Fault WB1[30].25'; 986 '~S001R03 Sealer Ctrlr 2 Required Rezeroing WB1[30].26'; 987 '~S001R03 Mig Barrel Replacement Warning WB1[30].27'; 988 '~S001R03 Mig Barrel Replacement Required WB1[30].28'; 989 '~S001R03 In Touch Up Mode WB1[30].29'; 990 '~S001R03 Touch Up Mode Not Enabled WB1[30].30'; 991 '~Spare WB1[30].31'; 992 '~S001R03 Laser Controller Fault WB1[31].0'; 993 '~S001R03 Laser Dirty Glass Warning WB1[31].1'; 994 '~S001R03 Laser Warning WB1[31].2'; 995 '~Spare WB1[31].3'; 996 '~Spare WB1[31].4'; 997 '~Spare WB1[31].5'; 998 '~Spare WB1[31].6'; 999 '~Spare WB1[31].7'; 1000 '~Spare WB1[31].8'; 1001 '~Spare WB1[31].9'; 1002 '~Spare WB1[31].10'; 1003 '~Spare WB1[31].11'; 1004 '~Spare WB1[31].12'; 1005 '~Spare WB1[31].13'; 1006 '~Spare WB1[31].14'; 1007 '~Spare WB1[31].15'; 1008 '~Spare WB1[31].16'; 1009 '~Spare WB1[31].17'; 1010 '~Spare WB1[31].18'; 1011 '~Spare WB1[31].19'; 1012 '~Spare WB1[31].20'; 1013 '~Spare WB1[31].21'; 1014 '~Spare WB1[31].22'; 1015 '~Spare WB1[31].23'; 1016 '~Spare WB1[31].24'; 1017 '~Spare WB1[31].25'; 1018 '~Spare WB1[31].26'; 1019 '~Spare WB1[31].27'; 1020 '~Spare WB1[31].28'; 1021 '~Spare WB1[31].29'; 1022 '~Spare WB1[31].30'; 1023 '~Spare WB1[31].31'; 1024 '~Spare WB1[32].0'; 1025 '~Spare WB1[32].1'; 1026 '~Spare WB1[32].2'; 1027 '~Spare WB1[32].3'; 1028 '~Spare WB1[32].4'; 1029 '~Spare WB1[32].5'; 1030 '~Spare WB1[32].6'; 1031 '~Spare WB1[32].7'; 1032 '~Spare WB1[32].8'; 1033 '~Spare WB1[32].9'; 1034 '~Spare WB1[32].10'; 1035 '~Spare WB1[32].11'; 1036 '~Spare WB1[32].12'; 1037 '~Spare WB1[32].13'; 1038 '~Spare WB1[32].14'; 1039 '~Spare WB1[32].15'; 1040 '~Spare WB1[32].16'; 1041 '~Spare WB1[32].17'; 1042 '~Spare WB1[32].18'; 1043 '~Spare WB1[32].19'; 1044 '~Spare WB1[32].20'; 1045 '~Spare WB1[32].21'; 1046 '~Spare WB1[32].22'; 1047 '~Spare WB1[32].23'; 1048 '~Spare WB1[32].24'; 1049 '~Spare WB1[32].25'; 1050 '~Spare WB1[32].26'; 1051 '~Spare WB1[32].27'; 1052 '~Spare WB1[32].28'; 1053 '~Spare WB1[32].29'; 1054 '~Spare WB1[32].30'; 1055 '~Spare WB1[32].31'; 1056 '~Spare WB1[33].0'; 1057 '~Spare WB1[33].1'; 1058 '~Spare WB1[33].2'; 1059 '~Spare WB1[33].3'; 1060 '~Spare WB1[33].4'; 1061 '~Spare WB1[33].5'; 1062 '~Spare WB1[33].6'; 1063 '~Spare WB1[33].7'; 1064 '~Spare WB1[33].8'; 1065 '~Spare WB1[33].9'; 1066 '~Spare WB1[33].10'; 1067 '~Spare WB1[33].11'; 1068 '~Spare WB1[33].12'; 1069 '~Spare WB1[33].13'; 1070 '~Spare WB1[33].14'; 1071 '~Spare WB1[33].15'; 1072 '~Spare WB1[33].16'; 1073 '~Spare WB1[33].17'; 1074 '~Spare WB1[33].18'; 1075 '~Spare WB1[33].19'; 1076 '~Spare WB1[33].20'; 1077 '~Spare WB1[33].21'; 1078 '~Spare WB1[33].22'; 1079 '~Spare WB1[33].23'; 1080 '~Spare WB1[33].24'; 1081 '~Spare WB1[33].25'; 1082 '~Spare WB1[33].26'; 1083 '~Spare WB1[33].27'; 1084 '~Spare WB1[33].28'; 1085 '~Spare WB1[33].29'; 1086 '~Spare WB1[33].30'; 1087 '~Spare WB1[33].31'; 1088 '~S001R04 Waiting Zone #1 Not Clear WB1[34].0'; 1089 '~S001R04 Waiting Zone #2 Not Clear WB1[34].1'; 1090 '~S001R04 Waiting Zone #3 Not Clear WB1[34].2'; 1091 '~S001R04 Waiting Zone #4 Not Clear WB1[34].3'; 1092 '~S001R04 Waiting Zone #5 Not Clear WB1[34].4'; 1093 '~S001R04 Waiting Zone #6 Not Clear WB1[34].5'; 1094 '~S001R04 Waiting Zone #7 Not Clear WB1[34].6'; 1095 '~S001R04 Waiting Zone #8 Not Clear WB1[34].7'; 1096 '~S001R04 Waiting Zone #9 Not Clear WB1[34].8'; 1097 '~S001R04 Waiting Zone #10 Not Clear WB1[34].9'; 1098 '~S001R04 Waiting Zone #11 Not Clear WB1[34].10'; 1099 '~S001R04 Waiting Zone #12 Not Clear WB1[34].11'; 1100 '~S001R04 Waiting Zone #13 Not Clear WB1[34].12'; 1101 '~S001R04 Waiting Zone #14 Not Clear WB1[34].13'; 1102 '~S001R04 Waiting Tip Dress Zone #1 Not Clear WB1[34].14'; 1103 '~S001R04 Waiting Tip Dress Zone #2 Not Clear WB1[34].15'; 1104 '~S001R04 Adjacent Robot xx-xx In Teach WB1[34].16'; 1105 '~S001R04 Adjacent Robot xx-xx In Teach WB1[34].17'; 1106 '~S001R04 Adjacent Robot xx-xx In Teach WB1[34].18'; 1107 '~S001R04 Adjacent Robot xx-xx In Teach WB1[34].19'; 1108 '~S001R04 Adjacent Robot xx-xx In Teach WB1[34].20'; 1109 '~S001R04 Adjacent Robot xx-xx In Teach WB1[34].21'; 1110 '~S001R04 Adjacent Robot xx-xx In Teach WB1[34].22'; 1111 '~S001R04 Adjacent Robot xx-xx In Teach WB1[34].23'; 1112 '~S001R04 Adjacent Robot xx-xx In Teach WB1[34].24'; 1113 '~S001R04 Adjacent Robot xx-xx In Teach WB1[34].25'; 1114 '~Spare WB1[34].26'; 1115 '~Spare WB1[34].27'; 1116 '~Spare WB1[34].28'; 1117 '~S001R04 Robot Not Clear Of Fixture WB1[34].29'; 1118 '~Spare WB1[34].30'; 1119 '~Spare WB1[34].31'; 1120 '~Spare WB1[35].0'; 1121 '~Spare WB1[35].1'; 1122 '~Spare WB1[35].2'; 1123 '~Spare WB1[35].3'; 1124 '~Spare WB1[35].4'; 1125 '~Spare WB1[35].5'; 1126 '~Spare WB1[35].6'; 1127 '~Spare WB1[35].7'; 1128 '~Spare WB1[35].8'; 1129 '~Spare WB1[35].9'; 1130 '~Spare WB1[35].10'; 1131 '~Spare WB1[35].11'; 1132 '~Spare WB1[35].12'; 1133 '~Spare WB1[35].13'; 1134 '~Spare WB1[35].14'; 1135 '~Spare WB1[35].15'; 1136 '~Spare WB1[35].16'; 1137 '~Spare WB1[35].17'; 1138 '~Spare WB1[35].18'; 1139 '~Spare WB1[35].19'; 1140 '~Spare WB1[35].20'; 1141 '~Spare WB1[35].21'; 1142 '~Spare WB1[35].22'; 1143 '~Spare WB1[35].23'; 1144 '~Spare WB1[35].24'; 1145 '~Spare WB1[35].25'; 1146 '~Spare WB1[35].26'; 1147 '~Spare WB1[35].27'; 1148 '~Spare WB1[35].28'; 1149 '~Spare WB1[35].29'; 1150 '~Spare WB1[35].30'; 1151 '~Spare WB1[35].31'; 1152 '~S001R04 Cycle Overtime WB1[36].0'; 1153 '~S001R04 In Bypass WB1[36].1'; 1154 '~S001R04 Battery Low WB1[36].2'; 1155 '~S001R04 Servo Over Torque WB1[36].3'; 1156 '~S001R04 Process Retry In Progress WB1[36].4'; 1157 '~Spare WB1[36].5'; 1158 '~S001R04 Robot Edit Occurred Ext App WB1[36].6'; 1159 '~S001R04 Robot Input Simmed WB1[36].7'; 1160 '~S001R04 Robot Output Simmed WB1[36].8'; 1161 '~Spare WB1[36].9'; 1162 '~Spare WB1[36].10'; 1163 '~Spare WB1[36].11'; 1164 '~Spare WB1[36].12'; 1165 '~Spare WB1[36].13'; 1166 '~Spare WB1[36].14'; 1167 '~Spare WB1[36].15'; 1168 '~S001R04F1B1.M.ModuleFlt - Externa App 1 I/O Module Warning WB1[36].16'; 1169 '~S001R04F2B1.M.ModuleFlt - Externa App 2 I/O Module Warning WB1[36].17'; 1170 '~S001R04F3B1.M.ModuleFlt - Externa App 3 I/O Module Warning WB1[36].18'; 1171 '~Spare WB1[36].19'; 1172 '~Spare WB1[36].20'; 1173 '~Spare WB1[36].21'; 1174 '~Spare WB1[36].22'; 1175 '~Spare WB1[36].23'; 1176 '~S001R04ES1 - S001R04 EtherNet Switch Port At Half Duplex WB1[36].24'; 1177 '~S001R04ES1 - S001R04 EtherNet Switch Config Changes Not Saved WB1[36].25'; 1178 '~S001R04ES1 - S001R04 EtherNet Switch Configuration Changed WB1[36].26'; 1179 '~S001R04ES1 - S001R04 EtherNet Switch Port With Excessive Errors WB1[36].27'; 1180 '~S001R04ES1 - S001R04 EtherNet Switch Port With Utilization Warning WB1[36].28'; 1181 '~S001R04ES1 - S001R04 EtherNet Switch Changes Require Reboot WB1[36].29'; 1182 '~Spare WB1[36].30'; 1183 '~Spare WB1[36].31'; 1184 '~Spare WB1[37].0'; 1185 '~Spare WB1[37].1'; 1186 '~S001R04 Servo Gun Tip Calib Request 1 WB1[37].2'; 1187 '~S001R04 I-Available Warning 1 WB1[37].3'; 1188 '~S001R04 Tip Dress Motor 1 Fault Bypassed WB1[37].4'; 1189 '~S001R04 Tip Change Notice 1 WB1[37].5'; 1190 '~S001R04 Bypass Tip Dresser 1 Selected WB1[37].6'; 1191 '~S001R04 Auto Tip Changer Low 1 WB1[37].7'; 1192 '~S001R04 Auto Tip Changer Empty 1 WB1[37].8'; 1193 '~S001R04 Tip Wear Ratio Warning 1 - Touch Up Tip Dress Program WB1[37].9'; 1194 '~S001R04 Stud Weld 1 Maintenance Reqd WB1[37].10'; 1195 '~S001R04 Stud Weld 1 Low Stud Warning WB1[37].11'; 1196 '~Spare WB1[37].12'; 1197 '~S001R04 Rivet 1 Low Rivet Warning WB1[37].13'; 1198 '~S001R04 Rivet 1 - Skip Once Initiated from Robot TP WB1[37].14'; 1199 '~S001R04 Rivet 1 - Skip Remaining Initiated from Robot TP WB1[37].15'; 1200 '~S001R04 Rivet 1 Preventive Maintenace Required WB1[37].16'; 1201 '~S001R04 Rivet 1 Magazine Low WB1[37].17'; 1202 '~S001R04 Tip Change 1 Bypassed WB1[37].18'; 1203 '~S001R04 Mig Weld Fluid Level Low WB1[37].19'; 1204 '~S001R04 Weld Ctrlr 1 Adaptive Mode Is Disabled WB1[37].20'; 1205 '~S001R04 Tip Cutter 1 Warning WB1[37].21'; 1206 '~S001R04 Rivet 1 Tape-Cut Required WB1[37].22'; 1207 '~S001R04 Wire Feeder Motor Over Current WB1[37].23'; 1208 '~Spare WB1[37].24'; 1209 '~S001R04 Sealer Ctrlr 1 Minor Fault WB1[37].25'; 1210 '~S001R04 Sealer Ctrlr 1 Required Rezeroing WB1[37].26'; 1211 '~S001R04 Loaded To Average WB1[37].27'; 1212 '~S001R04 Vision Process Aborted WB1[37].28'; 1213 '~S001R04 Vision System Trending WB1[37].29'; 1214 '~S001R04 Vision Out Of Tolerance WB1[37].30'; 1215 '~Spare WB1[37].31'; 1216 '~Spare WB1[38].0'; 1217 '~Spare WB1[38].1'; 1218 '~S001R04 Servo Gun Tip Calib Request 2 WB1[38].2'; 1219 '~S001R04 I-Available Warning 2 WB1[38].3'; 1220 '~S001R04 Tip Dress Motor 2 Fault Bypassed WB1[38].4'; 1221 '~S001R04 Tip Change Notice 2 WB1[38].5'; 1222 '~S001R04 Bypass Tip Dresser 2 Selected WB1[38].6'; 1223 '~S001R04 Auto Tip Changer Low 2 WB1[38].7'; 1224 '~S001R04 Auto Tip Changer Empty 2 WB1[38].8'; 1225 '~S001R04 Tip Wear Ratio Warning 2 - Touch Up Tip Dress Program WB1[38].9'; 1226 '~S001R04 Stud Weld 2 Maintenance Reqd WB1[38].10'; 1227 '~S001R04 Stud Weld 2 Low Stud Warning WB1[38].11'; 1228 '~Spare WB1[38].12'; 1229 '~S001R04 Rivet 2 Low Rivet Warning WB1[38].13'; 1230 '~S001R04 Rivet 2 - Skip Once Initiated from Robot TP WB1[38].14'; 1231 '~S001R04 Rivet 2 - Skip Remaining Initiated from Robot TP WB1[38].15'; 1232 '~S001R04 Rivet 2 Preventive Maintenace Required WB1[38].16'; 1233 '~S001R04 Rivet 2 Magazine Low WB1[38].17'; 1234 '~S001R04 Tip Change 2 Bypassed WB1[38].18'; 1235 '~S001R04 Laser Dirty Glass Warning WB1[38].19'; 1236 '~S001R04 Weld Ctrlr 2 Adaptive Mode Is Disabled WB1[38].20'; 1237 '~S001R04 Tip Cutter 2 Warning WB1[38].21'; 1238 '~S001R04 Rivet 2 Tape-Cut Required WB1[38].22'; 1239 '~S001R04 Mig Tip Nozzel Replacement Warning WB1[38].23'; 1240 '~S001R04 Mig Tip Nozzel Replacement Required WB1[38].24'; 1241 '~S001R04 Sealer Ctrlr 2 Minor Fault WB1[38].25'; 1242 '~S001R04 Sealer Ctrlr 2 Required Rezeroing WB1[38].26'; 1243 '~S001R04 Mig Barrel Replacement Warning WB1[38].27'; 1244 '~S001R04 Mig Barrel Replacement Required WB1[38].28'; 1245 '~S001R04 In Touch Up Mode WB1[38].29'; 1246 '~S001R04 Touch Up Mode Not Enabled WB1[38].30'; 1247 '~Spare WB1[38].31'; 1248 '~S001R04 Laser Controller Fault WB1[39].0'; 1249 '~S001R04 Laser Dirty Glass Warning WB1[39].1'; 1250 '~S001R04 Laser Warning WB1[39].2'; 1251 '~Spare WB1[39].3'; 1252 '~Spare WB1[39].4'; 1253 '~Spare WB1[39].5'; 1254 '~Spare WB1[39].6'; 1255 '~Spare WB1[39].7'; 1256 '~Spare WB1[39].8'; 1257 '~Spare WB1[39].9'; 1258 '~Spare WB1[39].10'; 1259 '~Spare WB1[39].11'; 1260 '~Spare WB1[39].12'; 1261 '~Spare WB1[39].13'; 1262 '~Spare WB1[39].14'; 1263 '~Spare WB1[39].15'; 1264 '~Spare WB1[39].16'; 1265 '~Spare WB1[39].17'; 1266 '~Spare WB1[39].18'; 1267 '~Spare WB1[39].19'; 1268 '~Spare WB1[39].20'; 1269 '~Spare WB1[39].21'; 1270 '~Spare WB1[39].22'; 1271 '~Spare WB1[39].23'; 1272 '~Spare WB1[39].24'; 1273 '~Spare WB1[39].25'; 1274 '~Spare WB1[39].26'; 1275 '~Spare WB1[39].27'; 1276 '~Spare WB1[39].28'; 1277 '~Spare WB1[39].29'; 1278 '~Spare WB1[39].30'; 1279 '~Spare WB1[39].31'; 1280 '~Spare WB1[40].0'; 1281 '~Spare WB1[40].1'; 1282 '~Spare WB1[40].2'; 1283 '~Spare WB1[40].3'; 1284 '~Spare WB1[40].4'; 1285 '~Spare WB1[40].5'; 1286 '~Spare WB1[40].6'; 1287 '~Spare WB1[40].7'; 1288 '~Spare WB1[40].8'; 1289 '~Spare WB1[40].9'; 1290 '~Spare WB1[40].10'; 1291 '~Spare WB1[40].11'; 1292 '~Spare WB1[40].12'; 1293 '~Spare WB1[40].13'; 1294 '~Spare WB1[40].14'; 1295 '~Spare WB1[40].15'; 1296 '~Spare WB1[40].16'; 1297 '~Spare WB1[40].17'; 1298 '~Spare WB1[40].18'; 1299 '~Spare WB1[40].19'; 1300 '~Spare WB1[40].20'; 1301 '~Spare WB1[40].21'; 1302 '~Spare WB1[40].22'; 1303 '~Spare WB1[40].23'; 1304 '~Spare WB1[40].24'; 1305 '~Spare WB1[40].25'; 1306 '~Spare WB1[40].26'; 1307 '~Spare WB1[40].27'; 1308 '~Spare WB1[40].28'; 1309 '~Spare WB1[40].29'; 1310 '~Spare WB1[40].30'; 1311 '~Spare WB1[40].31'; 1312 '~Spare WB1[41].0'; 1313 '~Spare WB1[41].1'; 1314 '~Spare WB1[41].2'; 1315 '~Spare WB1[41].3'; 1316 '~Spare WB1[41].4'; 1317 '~Spare WB1[41].5'; 1318 '~Spare WB1[41].6'; 1319 '~Spare WB1[41].7'; 1320 '~Spare WB1[41].8'; 1321 '~Spare WB1[41].9'; 1322 '~Spare WB1[41].10'; 1323 '~Spare WB1[41].11'; 1324 '~Spare WB1[41].12'; 1325 '~Spare WB1[41].13'; 1326 '~Spare WB1[41].14'; 1327 '~Spare WB1[41].15'; 1328 '~Spare WB1[41].16'; 1329 '~Spare WB1[41].17'; 1330 '~Spare WB1[41].18'; 1331 '~Spare WB1[41].19'; 1332 '~Spare WB1[41].20'; 1333 '~Spare WB1[41].21'; 1334 '~Spare WB1[41].22'; 1335 '~Spare WB1[41].23'; 1336 '~Spare WB1[41].24'; 1337 '~Spare WB1[41].25'; 1338 '~Spare WB1[41].26'; 1339 '~Spare WB1[41].27'; 1340 '~Spare WB1[41].28'; 1341 '~Spare WB1[41].29'; 1342 '~Spare WB1[41].30'; 1343 '~Spare WB1[41].31'; 1344 '~S001R05 Waiting Zone #1 Not Clear WB1[42].0'; 1345 '~S001R05 Waiting Zone #2 Not Clear WB1[42].1'; 1346 '~S001R05 Waiting Zone #3 Not Clear WB1[42].2'; 1347 '~S001R05 Waiting Zone #4 Not Clear WB1[42].3'; 1348 '~S001R05 Waiting Zone #5 Not Clear WB1[42].4'; 1349 '~S001R05 Waiting Zone #6 Not Clear WB1[42].5'; 1350 '~S001R05 Waiting Zone #7 Not Clear WB1[42].6'; 1351 '~S001R05 Waiting Zone #8 Not Clear WB1[42].7'; 1352 '~S001R05 Waiting Zone #9 Not Clear WB1[42].8'; 1353 '~S001R05 Waiting Zone #10 Not Clear WB1[42].9'; 1354 '~S001R05 Waiting Zone #11 Not Clear WB1[42].10'; 1355 '~S001R05 Waiting Zone #12 Not Clear WB1[42].11'; 1356 '~S001R05 Waiting Zone #13 Not Clear WB1[42].12'; 1357 '~S001R05 Waiting Zone #14 Not Clear WB1[42].13'; 1358 '~S001R05 Waiting Tip Dress Zone #1 Not Clear WB1[42].14'; 1359 '~S001R05 Waiting Tip Dress Zone #2 Not Clear WB1[42].15'; 1360 '~S001R05 Adjacent Robot xx-xx In Teach WB1[42].16'; 1361 '~S001R05 Adjacent Robot xx-xx In Teach WB1[42].17'; 1362 '~S001R05 Adjacent Robot xx-xx In Teach WB1[42].18'; 1363 '~S001R05 Adjacent Robot xx-xx In Teach WB1[42].19'; 1364 '~S001R05 Adjacent Robot xx-xx In Teach WB1[42].20'; 1365 '~S001R05 Adjacent Robot xx-xx In Teach WB1[42].21'; 1366 '~S001R05 Adjacent Robot xx-xx In Teach WB1[42].22'; 1367 '~S001R05 Adjacent Robot xx-xx In Teach WB1[42].23'; 1368 '~S001R05 Adjacent Robot xx-xx In Teach WB1[42].24'; 1369 '~S001R05 Adjacent Robot xx-xx In Teach WB1[42].25'; 1370 '~Spare WB1[42].26'; 1371 '~Spare WB1[42].27'; 1372 '~Spare WB1[42].28'; 1373 '~S001R05 Robot Not Clear Of Fixture WB1[42].29'; 1374 '~Spare WB1[42].30'; 1375 '~Spare WB1[42].31'; 1376 '~Spare WB1[43].0'; 1377 '~Spare WB1[43].1'; 1378 '~Spare WB1[43].2'; 1379 '~Spare WB1[43].3'; 1380 '~Spare WB1[43].4'; 1381 '~Spare WB1[43].5'; 1382 '~Spare WB1[43].6'; 1383 '~Spare WB1[43].7'; 1384 '~Spare WB1[43].8'; 1385 '~Spare WB1[43].9'; 1386 '~Spare WB1[43].10'; 1387 '~Spare WB1[43].11'; 1388 '~Spare WB1[43].12'; 1389 '~Spare WB1[43].13'; 1390 '~Spare WB1[43].14'; 1391 '~Spare WB1[43].15'; 1392 '~Spare WB1[43].16'; 1393 '~Spare WB1[43].17'; 1394 '~Spare WB1[43].18'; 1395 '~Spare WB1[43].19'; 1396 '~Spare WB1[43].20'; 1397 '~Spare WB1[43].21'; 1398 '~Spare WB1[43].22'; 1399 '~Spare WB1[43].23'; 1400 '~Spare WB1[43].24'; 1401 '~Spare WB1[43].25'; 1402 '~Spare WB1[43].26'; 1403 '~Spare WB1[43].27'; 1404 '~Spare WB1[43].28'; 1405 '~Spare WB1[43].29'; 1406 '~Spare WB1[43].30'; 1407 '~Spare WB1[43].31'; 1408 '~S001R05 Cycle Overtime WB1[44].0'; 1409 '~S001R05 In Bypass WB1[44].1'; 1410 '~S001R05 Battery Low WB1[44].2'; 1411 '~S001R05 Servo Over Torque WB1[44].3'; 1412 '~S001R05 Process Retry In Progress WB1[44].4'; 1413 '~Spare WB1[44].5'; 1414 '~S001R05 Robot Edit Occurred Ext App WB1[44].6'; 1415 '~S001R05 Robot Input Simmed WB1[44].7'; 1416 '~S001R05 Robot Output Simmed WB1[44].8'; 1417 '~Spare WB1[44].9'; 1418 '~Spare WB1[44].10'; 1419 '~Spare WB1[44].11'; 1420 '~Spare WB1[44].12'; 1421 '~Spare WB1[44].13'; 1422 '~Spare WB1[44].14'; 1423 '~Spare WB1[44].15'; 1424 '~S001R05F1B1.M.ModuleFlt - Externa App 1 I/O Module Warning WB1[44].16'; 1425 '~S001R05F2B1.M.ModuleFlt - Externa App 2 I/O Module Warning WB1[44].17'; 1426 '~S001R05F3B1.M.ModuleFlt - Externa App 3 I/O Module Warning WB1[44].18'; 1427 '~Spare WB1[44].19'; 1428 '~Spare WB1[44].20'; 1429 '~Spare WB1[44].21'; 1430 '~Spare WB1[44].22'; 1431 '~Spare WB1[44].23'; 1432 '~S001R05ES1 - S001R05 EtherNet Switch Port At Half Duplex WB1[44].24'; 1433 '~S001R05ES1 - S001R05 EtherNet Switch Config Changes Not Saved WB1[44].25'; 1434 '~S001R05ES1 - S001R05 EtherNet Switch Configuration Changed WB1[44].26'; 1435 '~S001R05ES1 - S001R05 EtherNet Switch Port With Excessive Errors WB1[44].27'; 1436 '~S001R05ES1 - S001R05 EtherNet Switch Port With Utilization Warning WB1[44].28'; 1437 '~S001R05ES1 - S001R05 EtherNet Switch Changes Require Reboot WB1[44].29'; 1438 '~Spare WB1[44].30'; 1439 '~Spare WB1[44].31'; 1440 '~Spare WB1[45].0'; 1441 '~Spare WB1[45].1'; 1442 '~S001R05 Servo Gun Tip Calib Request 1 WB1[45].2'; 1443 '~S001R05 I-Available Warning 1 WB1[45].3'; 1444 '~S001R05 Tip Dress Motor 1 Fault Bypassed WB1[45].4'; 1445 '~S001R05 Tip Change Notice 1 WB1[45].5'; 1446 '~S001R05 Bypass Tip Dresser 1 Selected WB1[45].6'; 1447 '~S001R05 Auto Tip Changer Low 1 WB1[45].7'; 1448 '~S001R05 Auto Tip Changer Empty 1 WB1[45].8'; 1449 '~S001R05 Tip Wear Ratio Warning 1 - Touch Up Tip Dress Program WB1[45].9'; 1450 '~S001R05 Stud Weld 1 Maintenance Reqd WB1[45].10'; 1451 '~S001R05 Stud Weld 1 Low Stud Warning WB1[45].11'; 1452 '~Spare WB1[45].12'; 1453 '~S001R05 Rivet 1 Low Rivet Warning WB1[45].13'; 1454 '~S001R05 Rivet 1 - Skip Once Initiated from Robot TP WB1[45].14'; 1455 '~S001R05 Rivet 1 - Skip Remaining Initiated from Robot TP WB1[45].15'; 1456 '~S001R05 Rivet 1 Preventive Maintenace Required WB1[45].16'; 1457 '~S001R05 Rivet 1 Magazine Low WB1[45].17'; 1458 '~S001R05 Tip Change 1 Bypassed WB1[45].18'; 1459 '~S001R05 Mig Weld Fluid Level Low WB1[45].19'; 1460 '~S001R05 Weld Ctrlr 1 Adaptive Mode Is Disabled WB1[45].20'; 1461 '~S001R05 Tip Cutter 1 Warning WB1[45].21'; 1462 '~S001R05 Rivet 1 Tape-Cut Required WB1[45].22'; 1463 '~S001R05 Wire Feeder Motor Over Current WB1[45].23'; 1464 '~Spare WB1[45].24'; 1465 '~S001R05 Sealer Ctrlr 1 Minor Fault WB1[45].25'; 1466 '~S001R05 Sealer Ctrlr 1 Required Rezeroing WB1[45].26'; 1467 '~S001R05 Loaded To Average WB1[45].27'; 1468 '~S001R05 Vision Process Aborted WB1[45].28'; 1469 '~S001R05 Vision System Trending WB1[45].29'; 1470 '~S001R05 Vision Out Of Tolerance WB1[45].30'; 1471 '~Spare WB1[45].31'; 1472 '~Spare WB1[46].0'; 1473 '~Spare WB1[46].1'; 1474 '~S001R05 Servo Gun Tip Calib Request 2 WB1[46].2'; 1475 '~S001R05 I-Available Warning 2 WB1[46].3'; 1476 '~S001R05 Tip Dress Motor 2 Fault Bypassed WB1[46].4'; 1477 '~S001R05 Tip Change Notice 2 WB1[46].5'; 1478 '~S001R05 Bypass Tip Dresser 2 Selected WB1[46].6'; 1479 '~S001R05 Auto Tip Changer Low 2 WB1[46].7'; 1480 '~S001R05 Auto Tip Changer Empty 2 WB1[46].8'; 1481 '~S001R05 Tip Wear Ratio Warning 2 - Touch Up Tip Dress Program WB1[46].9'; 1482 '~S001R05 Stud Weld 2 Maintenance Reqd WB1[46].10'; 1483 '~S001R05 Stud Weld 2 Low Stud Warning WB1[46].11'; 1484 '~Spare WB1[46].12'; 1485 '~S001R05 Rivet 2 Low Rivet Warning WB1[46].13'; 1486 '~S001R05 Rivet 2 - Skip Once Initiated from Robot TP WB1[46].14'; 1487 '~S001R05 Rivet 2 - Skip Remaining Initiated from Robot TP WB1[46].15'; 1488 '~S001R05 Rivet 2 Preventive Maintenace Required WB1[46].16'; 1489 '~S001R05 Rivet 2 Magazine Low WB1[46].17'; 1490 '~S001R05 Tip Change 2 Bypassed WB1[46].18'; 1491 '~S001R05 Laser Dirty Glass Warning WB1[46].19'; 1492 '~S001R05 Weld Ctrlr 2 Adaptive Mode Is Disabled WB1[46].20'; 1493 '~S001R05 Tip Cutter 2 Warning WB1[46].21'; 1494 '~S001R05 Rivet 2 Tape-Cut Required WB1[46].22'; 1495 '~S001R05 Mig Tip Nozzel Replacement Warning WB1[46].23'; 1496 '~S001R05 Mig Tip Nozzel Replacement Required WB1[46].24'; 1497 '~S001R05 Sealer Ctrlr 2 Minor Fault WB1[46].25'; 1498 '~S001R05 Sealer Ctrlr 2 Required Rezeroing WB1[46].26'; 1499 '~S001R05 Mig Barrel Replacement Warning WB1[46].27'; 1500 '~S001R05 Mig Barrel Replacement Required WB1[46].28'; 1501 '~S001R05 In Touch Up Mode WB1[46].29'; 1502 '~S001R05 Touch Up Mode Not Enabled WB1[46].30'; 1503 '~Spare WB1[46].31'; 1504 '~S001R05 Laser Controller Fault WB1[47].0'; 1505 '~S001R05 Laser Dirty Glass Warning WB1[47].1'; 1506 '~S001R05 Laser Warning WB1[47].2'; 1507 '~Spare WB1[47].3'; 1508 '~Spare WB1[47].4'; 1509 '~Spare WB1[47].5'; 1510 '~Spare WB1[47].6'; 1511 '~Spare WB1[47].7'; 1512 '~Spare WB1[47].8'; 1513 '~Spare WB1[47].9'; 1514 '~Spare WB1[47].10'; 1515 '~Spare WB1[47].11'; 1516 '~Spare WB1[47].12'; 1517 '~Spare WB1[47].13'; 1518 '~Spare WB1[47].14'; 1519 '~Spare WB1[47].15'; 1520 '~Spare WB1[47].16'; 1521 '~Spare WB1[47].17'; 1522 '~Spare WB1[47].18'; 1523 '~Spare WB1[47].19'; 1524 '~Spare WB1[47].20'; 1525 '~Spare WB1[47].21'; 1526 '~Spare WB1[47].22'; 1527 '~Spare WB1[47].23'; 1528 '~Spare WB1[47].24'; 1529 '~Spare WB1[47].25'; 1530 '~Spare WB1[47].26'; 1531 '~Spare WB1[47].27'; 1532 '~Spare WB1[47].28'; 1533 '~Spare WB1[47].29'; 1534 '~Spare WB1[47].30'; 1535 '~Spare WB1[47].31'; 1536 '~Spare WB1[48].0'; 1537 '~Spare WB1[48].1'; 1538 '~Spare WB1[48].2'; 1539 '~Spare WB1[48].3'; 1540 '~Spare WB1[48].4'; 1541 '~Spare WB1[48].5'; 1542 '~Spare WB1[48].6'; 1543 '~Spare WB1[48].7'; 1544 '~Spare WB1[48].8'; 1545 '~Spare WB1[48].9'; 1546 '~Spare WB1[48].10'; 1547 '~Spare WB1[48].11'; 1548 '~Spare WB1[48].12'; 1549 '~Spare WB1[48].13'; 1550 '~Spare WB1[48].14'; 1551 '~Spare WB1[48].15'; 1552 '~Spare WB1[48].16'; 1553 '~Spare WB1[48].17'; 1554 '~Spare WB1[48].18'; 1555 '~Spare WB1[48].19'; 1556 '~Spare WB1[48].20'; 1557 '~Spare WB1[48].21'; 1558 '~Spare WB1[48].22'; 1559 '~Spare WB1[48].23'; 1560 '~Spare WB1[48].24'; 1561 '~Spare WB1[48].25'; 1562 '~Spare WB1[48].26'; 1563 '~Spare WB1[48].27'; 1564 '~Spare WB1[48].28'; 1565 '~Spare WB1[48].29'; 1566 '~Spare WB1[48].30'; 1567 '~Spare WB1[48].31'; 1568 '~Spare WB1[49].0'; 1569 '~Spare WB1[49].1'; 1570 '~Spare WB1[49].2'; 1571 '~Spare WB1[49].3'; 1572 '~Spare WB1[49].4'; 1573 '~Spare WB1[49].5'; 1574 '~Spare WB1[49].6'; 1575 '~Spare WB1[49].7'; 1576 '~Spare WB1[49].8'; 1577 '~Spare WB1[49].9'; 1578 '~Spare WB1[49].10'; 1579 '~Spare WB1[49].11'; 1580 '~Spare WB1[49].12'; 1581 '~Spare WB1[49].13'; 1582 '~Spare WB1[49].14'; 1583 '~Spare WB1[49].15'; 1584 '~Spare WB1[49].16'; 1585 '~Spare WB1[49].17'; 1586 '~Spare WB1[49].18'; 1587 '~Spare WB1[49].19'; 1588 '~Spare WB1[49].20'; 1589 '~Spare WB1[49].21'; 1590 '~Spare WB1[49].22'; 1591 '~Spare WB1[49].23'; 1592 '~Spare WB1[49].24'; 1593 '~Spare WB1[49].25'; 1594 '~Spare WB1[49].26'; 1595 '~Spare WB1[49].27'; 1596 '~Spare WB1[49].28'; 1597 '~Spare WB1[49].29'; 1598 '~Spare WB1[49].30'; 1599 '~Spare WB1[49].31'; 1600 '~S001R06 Waiting Zone #1 Not Clear WB1[50].0'; 1601 '~S001R06 Waiting Zone #2 Not Clear WB1[50].1'; 1602 '~S001R06 Waiting Zone #3 Not Clear WB1[50].2'; 1603 '~S001R06 Waiting Zone #4 Not Clear WB1[50].3'; 1604 '~S001R06 Waiting Zone #5 Not Clear WB1[50].4'; 1605 '~S001R06 Waiting Zone #6 Not Clear WB1[50].5'; 1606 '~S001R06 Waiting Zone #7 Not Clear WB1[50].6'; 1607 '~S001R06 Waiting Zone #8 Not Clear WB1[50].7'; 1608 '~S001R06 Waiting Zone #9 Not Clear WB1[50].8'; 1609 '~S001R06 Waiting Zone #10 Not Clear WB1[50].9'; 1610 '~S001R06 Waiting Zone #11 Not Clear WB1[50].10'; 1611 '~S001R06 Waiting Zone #12 Not Clear WB1[50].11'; 1612 '~S001R06 Waiting Zone #13 Not Clear WB1[50].12'; 1613 '~S001R06 Waiting Zone #14 Not Clear WB1[50].13'; 1614 '~S001R06 Waiting Tip Dress Zone #1 Not Clear WB1[50].14'; 1615 '~S001R06 Waiting Tip Dress Zone #2 Not Clear WB1[50].15'; 1616 '~S001R06 Adjacent Robot xx-xx In Teach WB1[50].16'; 1617 '~S001R06 Adjacent Robot xx-xx In Teach WB1[50].17'; 1618 '~S001R06 Adjacent Robot xx-xx In Teach WB1[50].18'; 1619 '~S001R06 Adjacent Robot xx-xx In Teach WB1[50].19'; 1620 '~S001R06 Adjacent Robot xx-xx In Teach WB1[50].20'; 1621 '~S001R06 Adjacent Robot xx-xx In Teach WB1[50].21'; 1622 '~S001R06 Adjacent Robot xx-xx In Teach WB1[50].22'; 1623 '~S001R06 Adjacent Robot xx-xx In Teach WB1[50].23'; 1624 '~S001R06 Adjacent Robot xx-xx In Teach WB1[50].24'; 1625 '~S001R06 Adjacent Robot xx-xx In Teach WB1[50].25'; 1626 '~Spare WB1[50].26'; 1627 '~Spare WB1[50].27'; 1628 '~Spare WB1[50].28'; 1629 '~S001R06 Robot Not Clear Of Fixture WB1[50].29'; 1630 '~Spare WB1[50].30'; 1631 '~Spare WB1[50].31'; 1632 '~Spare WB1[51].0'; 1633 '~Spare WB1[51].1'; 1634 '~Spare WB1[51].2'; 1635 '~Spare WB1[51].3'; 1636 '~Spare WB1[51].4'; 1637 '~Spare WB1[51].5'; 1638 '~Spare WB1[51].6'; 1639 '~Spare WB1[51].7'; 1640 '~Spare WB1[51].8'; 1641 '~Spare WB1[51].9'; 1642 '~Spare WB1[51].10'; 1643 '~Spare WB1[51].11'; 1644 '~Spare WB1[51].12'; 1645 '~Spare WB1[51].13'; 1646 '~Spare WB1[51].14'; 1647 '~Spare WB1[51].15'; 1648 '~Spare WB1[51].16'; 1649 '~Spare WB1[51].17'; 1650 '~Spare WB1[51].18'; 1651 '~Spare WB1[51].19'; 1652 '~Spare WB1[51].20'; 1653 '~Spare WB1[51].21'; 1654 '~Spare WB1[51].22'; 1655 '~Spare WB1[51].23'; 1656 '~Spare WB1[51].24'; 1657 '~Spare WB1[51].25'; 1658 '~Spare WB1[51].26'; 1659 '~Spare WB1[51].27'; 1660 '~Spare WB1[51].28'; 1661 '~Spare WB1[51].29'; 1662 '~Spare WB1[51].30'; 1663 '~Spare WB1[51].31'; 1664 '~S001R06 Cycle Overtime WB1[52].0'; 1665 '~S001R06 In Bypass WB1[52].1'; 1666 '~S001R06 Battery Low WB1[52].2'; 1667 '~S001R06 Servo Over Torque WB1[52].3'; 1668 '~S001R06 Process Retry In Progress WB1[52].4'; 1669 '~Spare WB1[52].5'; 1670 '~S001R06 Robot Edit Occurred Ext App WB1[52].6'; 1671 '~S001R06 Robot Input Simmed WB1[52].7'; 1672 '~S001R06 Robot Output Simmed WB1[52].8'; 1673 '~Spare WB1[52].9'; 1674 '~Spare WB1[52].10'; 1675 '~Spare WB1[52].11'; 1676 '~Spare WB1[52].12'; 1677 '~Spare WB1[52].13'; 1678 '~Spare WB1[52].14'; 1679 '~Spare WB1[52].15'; 1680 '~S001R06F1B1.M.ModuleFlt - Externa App 1 I/O Module Warning WB1[52].16'; 1681 '~S001R06F2B1.M.ModuleFlt - Externa App 2 I/O Module Warning WB1[52].17'; 1682 '~S001R06F3B1.M.ModuleFlt - Externa App 3 I/O Module Warning WB1[52].18'; 1683 '~Spare WB1[52].19'; 1684 '~Spare WB1[52].20'; 1685 '~Spare WB1[52].21'; 1686 '~Spare WB1[52].22'; 1687 '~Spare WB1[52].23'; 1688 '~S001R06ES1 - S001R06 EtherNet Switch Port At Half Duplex WB1[52].24'; 1689 '~S001R06ES1 - S001R06 EtherNet Switch Config Changes Not Saved WB1[52].25'; 1690 '~S001R06ES1 - S001R06 EtherNet Switch Configuration Changed WB1[52].26'; 1691 '~S001R06ES1 - S001R06 EtherNet Switch Port With Excessive Errors WB1[52].27'; 1692 '~S001R06ES1 - S001R06 EtherNet Switch Port With Utilization Warning WB1[52].28'; 1693 '~S001R06ES1 - S001R06 EtherNet Switch Changes Require Reboot WB1[52].29'; 1694 '~Spare WB1[52].30'; 1695 '~Spare WB1[52].31'; 1696 '~Spare WB1[53].0'; 1697 '~Spare WB1[53].1'; 1698 '~S001R06 Servo Gun Tip Calib Request 1 WB1[53].2'; 1699 '~S001R06 I-Available Warning 1 WB1[53].3'; 1700 '~S001R06 Tip Dress Motor 1 Fault Bypassed WB1[53].4'; 1701 '~S001R06 Tip Change Notice 1 WB1[53].5'; 1702 '~S001R06 Bypass Tip Dresser 1 Selected WB1[53].6'; 1703 '~S001R06 Auto Tip Changer Low 1 WB1[53].7'; 1704 '~S001R06 Auto Tip Changer Empty 1 WB1[53].8'; 1705 '~S001R06 Tip Wear Ratio Warning 1 - Touch Up Tip Dress Program WB1[53].9'; 1706 '~S001R06 Stud Weld 1 Maintenance Reqd WB1[53].10'; 1707 '~S001R06 Stud Weld 1 Low Stud Warning WB1[53].11'; 1708 '~Spare WB1[53].12'; 1709 '~S001R06 Rivet 1 Low Rivet Warning WB1[53].13'; 1710 '~S001R06 Rivet 1 - Skip Once Initiated from Robot TP WB1[53].14'; 1711 '~S001R06 Rivet 1 - Skip Remaining Initiated from Robot TP WB1[53].15'; 1712 '~S001R06 Rivet 1 Preventive Maintenace Required WB1[53].16'; 1713 '~S001R06 Rivet 1 Magazine Low WB1[53].17'; 1714 '~S001R06 Tip Change 1 Bypassed WB1[53].18'; 1715 '~S001R06 Mig Weld Fluid Level Low WB1[53].19'; 1716 '~S001R06 Weld Ctrlr 1 Adaptive Mode Is Disabled WB1[53].20'; 1717 '~S001R06 Tip Cutter 1 Warning WB1[53].21'; 1718 '~S001R06 Rivet 1 Tape-Cut Required WB1[53].22'; 1719 '~S001R06 Wire Feeder Motor Over Current WB1[53].23'; 1720 '~Spare WB1[53].24'; 1721 '~S001R06 Sealer Ctrlr 1 Minor Fault WB1[53].25'; 1722 '~S001R06 Sealer Ctrlr 1 Required Rezeroing WB1[53].26'; 1723 '~S001R06 Loaded To Average WB1[53].27'; 1724 '~S001R06 Vision Process Aborted WB1[53].28'; 1725 '~S001R06 Vision System Trending WB1[53].29'; 1726 '~S001R06 Vision Out Of Tolerance WB1[53].30'; 1727 '~Spare WB1[53].31'; 1728 '~Spare WB1[54].0'; 1729 '~Spare WB1[54].1'; 1730 '~S001R06 Servo Gun Tip Calib Request 2 WB1[54].2'; 1731 '~S001R06 I-Available Warning 2 WB1[54].3'; 1732 '~S001R06 Tip Dress Motor 2 Fault Bypassed WB1[54].4'; 1733 '~S001R06 Tip Change Notice 2 WB1[54].5'; 1734 '~S001R06 Bypass Tip Dresser 2 Selected WB1[54].6'; 1735 '~S001R06 Auto Tip Changer Low 2 WB1[54].7'; 1736 '~S001R06 Auto Tip Changer Empty 2 WB1[54].8'; 1737 '~S001R06 Tip Wear Ratio Warning 2 - Touch Up Tip Dress Program WB1[54].9'; 1738 '~S001R06 Stud Weld 2 Maintenance Reqd WB1[54].10'; 1739 '~S001R06 Stud Weld 2 Low Stud Warning WB1[54].11'; 1740 '~Spare WB1[54].12'; 1741 '~S001R06 Rivet 2 Low Rivet Warning WB1[54].13'; 1742 '~S001R06 Rivet 2 - Skip Once Initiated from Robot TP WB1[54].14'; 1743 '~S001R06 Rivet 2 - Skip Remaining Initiated from Robot TP WB1[54].15'; 1744 '~S001R06 Rivet 2 Preventive Maintenace Required WB1[54].16'; 1745 '~S001R06 Rivet 2 Magazine Low WB1[54].17'; 1746 '~S001R06 Tip Change 2 Bypassed WB1[54].18'; 1747 '~S001R06 Laser Dirty Glass Warning WB1[54].19'; 1748 '~S001R06 Weld Ctrlr 2 Adaptive Mode Is Disabled WB1[54].20'; 1749 '~S001R06 Tip Cutter 2 Warning WB1[54].21'; 1750 '~S001R06 Rivet 2 Tape-Cut Required WB1[54].22'; 1751 '~S001R06 Mig Tip Nozzel Replacement Warning WB1[54].23'; 1752 '~S001R06 Mig Tip Nozzel Replacement Required WB1[54].24'; 1753 '~S001R06 Sealer Ctrlr 2 Minor Fault WB1[54].25'; 1754 '~S001R06 Sealer Ctrlr 2 Required Rezeroing WB1[54].26'; 1755 '~S001R06 Mig Barrel Replacement Warning WB1[54].27'; 1756 '~S001R06 Mig Barrel Replacement Required WB1[54].28'; 1757 '~S001R06 In Touch Up Mode WB1[54].29'; 1758 '~S001R06 Touch Up Mode Not Enabled WB1[54].30'; 1759 '~Spare WB1[54].31'; 1760 '~S001R06 Laser Controller Fault WB1[55].0'; 1761 '~S001R06 Laser Dirty Glass Warning WB1[55].1'; 1762 '~S001R06 Laser Warning WB1[55].2'; 1763 '~Spare WB1[55].3'; 1764 '~Spare WB1[55].4'; 1765 '~Spare WB1[55].5'; 1766 '~Spare WB1[55].6'; 1767 '~Spare WB1[55].7'; 1768 '~Spare WB1[55].8'; 1769 '~Spare WB1[55].9'; 1770 '~Spare WB1[55].10'; 1771 '~Spare WB1[55].11'; 1772 '~Spare WB1[55].12'; 1773 '~Spare WB1[55].13'; 1774 '~Spare WB1[55].14'; 1775 '~Spare WB1[55].15'; 1776 '~Spare WB1[55].16'; 1777 '~Spare WB1[55].17'; 1778 '~Spare WB1[55].18'; 1779 '~Spare WB1[55].19'; 1780 '~Spare WB1[55].20'; 1781 '~Spare WB1[55].21'; 1782 '~Spare WB1[55].22'; 1783 '~Spare WB1[55].23'; 1784 '~Spare WB1[55].24'; 1785 '~Spare WB1[55].25'; 1786 '~Spare WB1[55].26'; 1787 '~Spare WB1[55].27'; 1788 '~Spare WB1[55].28'; 1789 '~Spare WB1[55].29'; 1790 '~Spare WB1[55].30'; 1791 '~Spare WB1[55].31'; 1792 '~Spare WB1[56].0'; 1793 '~Spare WB1[56].1'; 1794 '~Spare WB1[56].2'; 1795 '~Spare WB1[56].3'; 1796 '~Spare WB1[56].4'; 1797 '~Spare WB1[56].5'; 1798 '~Spare WB1[56].6'; 1799 '~Spare WB1[56].7'; 1800 '~Spare WB1[56].8'; 1801 '~Spare WB1[56].9'; 1802 '~Spare WB1[56].10'; 1803 '~Spare WB1[56].11'; 1804 '~Spare WB1[56].12'; 1805 '~Spare WB1[56].13'; 1806 '~Spare WB1[56].14'; 1807 '~Spare WB1[56].15'; 1808 '~Spare WB1[56].16'; 1809 '~Spare WB1[56].17'; 1810 '~Spare WB1[56].18'; 1811 '~Spare WB1[56].19'; 1812 '~Spare WB1[56].20'; 1813 '~Spare WB1[56].21'; 1814 '~Spare WB1[56].22'; 1815 '~Spare WB1[56].23'; 1816 '~Spare WB1[56].24'; 1817 '~Spare WB1[56].25'; 1818 '~Spare WB1[56].26'; 1819 '~Spare WB1[56].27'; 1820 '~Spare WB1[56].28'; 1821 '~Spare WB1[56].29'; 1822 '~Spare WB1[56].30'; 1823 '~Spare WB1[56].31'; 1824 '~Spare WB1[57].0'; 1825 '~Spare WB1[57].1'; 1826 '~Spare WB1[57].2'; 1827 '~Spare WB1[57].3'; 1828 '~Spare WB1[57].4'; 1829 '~Spare WB1[57].5'; 1830 '~Spare WB1[57].6'; 1831 '~Spare WB1[57].7'; 1832 '~Spare WB1[57].8'; 1833 '~Spare WB1[57].9'; 1834 '~Spare WB1[57].10'; 1835 '~Spare WB1[57].11'; 1836 '~Spare WB1[57].12'; 1837 '~Spare WB1[57].13'; 1838 '~Spare WB1[57].14'; 1839 '~Spare WB1[57].15'; 1840 '~Spare WB1[57].16'; 1841 '~Spare WB1[57].17'; 1842 '~Spare WB1[57].18'; 1843 '~Spare WB1[57].19'; 1844 '~Spare WB1[57].20'; 1845 '~Spare WB1[57].21'; 1846 '~Spare WB1[57].22'; 1847 '~Spare WB1[57].23'; 1848 '~Spare WB1[57].24'; 1849 '~Spare WB1[57].25'; 1850 '~Spare WB1[57].26'; 1851 '~Spare WB1[57].27'; 1852 '~Spare WB1[57].28'; 1853 '~Spare WB1[57].29'; 1854 '~Spare WB1[57].30'; 1855 '~Spare WB1[57].31'; 1856 '~S001R07 Waiting Zone #1 Not Clear WB1[58].0'; 1857 '~S001R07 Waiting Zone #2 Not Clear WB1[58].1'; 1858 '~S001R07 Waiting Zone #3 Not Clear WB1[58].2'; 1859 '~S001R07 Waiting Zone #4 Not Clear WB1[58].3'; 1860 '~S001R07 Waiting Zone #5 Not Clear WB1[58].4'; 1861 '~S001R07 Waiting Zone #6 Not Clear WB1[58].5'; 1862 '~S001R07 Waiting Zone #7 Not Clear WB1[58].6'; 1863 '~S001R07 Waiting Zone #8 Not Clear WB1[58].7'; 1864 '~S001R07 Waiting Zone #9 Not Clear WB1[58].8'; 1865 '~S001R07 Waiting Zone #10 Not Clear WB1[58].9'; 1866 '~S001R07 Waiting Zone #11 Not Clear WB1[58].10'; 1867 '~S001R07 Waiting Zone #12 Not Clear WB1[58].11'; 1868 '~S001R07 Waiting Zone #13 Not Clear WB1[58].12'; 1869 '~S001R07 Waiting Zone #14 Not Clear WB1[58].13'; 1870 '~S001R07 Waiting Tip Dress Zone #1 Not Clear WB1[58].14'; 1871 '~S001R07 Waiting Tip Dress Zone #2 Not Clear WB1[58].15'; 1872 '~S001R07 Adjacent Robot xx-xx In Teach WB1[58].16'; 1873 '~S001R07 Adjacent Robot xx-xx In Teach WB1[58].17'; 1874 '~S001R07 Adjacent Robot xx-xx In Teach WB1[58].18'; 1875 '~S001R07 Adjacent Robot xx-xx In Teach WB1[58].19'; 1876 '~S001R07 Adjacent Robot xx-xx In Teach WB1[58].20'; 1877 '~S001R07 Adjacent Robot xx-xx In Teach WB1[58].21'; 1878 '~S001R07 Adjacent Robot xx-xx In Teach WB1[58].22'; 1879 '~S001R07 Adjacent Robot xx-xx In Teach WB1[58].23'; 1880 '~S001R07 Adjacent Robot xx-xx In Teach WB1[58].24'; 1881 '~S001R07 Adjacent Robot xx-xx In Teach WB1[58].25'; 1882 '~Spare WB1[58].26'; 1883 '~Spare WB1[58].27'; 1884 '~Spare WB1[58].28'; 1885 '~S001R07 Robot Not Clear Of Fixture WB1[58].29'; 1886 '~Spare WB1[58].30'; 1887 '~Spare WB1[58].31'; 1888 '~Spare WB1[59].0'; 1889 '~Spare WB1[59].1'; 1890 '~Spare WB1[59].2'; 1891 '~Spare WB1[59].3'; 1892 '~Spare WB1[59].4'; 1893 '~Spare WB1[59].5'; 1894 '~Spare WB1[59].6'; 1895 '~Spare WB1[59].7'; 1896 '~Spare WB1[59].8'; 1897 '~Spare WB1[59].9'; 1898 '~Spare WB1[59].10'; 1899 '~Spare WB1[59].11'; 1900 '~Spare WB1[59].12'; 1901 '~Spare WB1[59].13'; 1902 '~Spare WB1[59].14'; 1903 '~Spare WB1[59].15'; 1904 '~Spare WB1[59].16'; 1905 '~Spare WB1[59].17'; 1906 '~Spare WB1[59].18'; 1907 '~Spare WB1[59].19'; 1908 '~Spare WB1[59].20'; 1909 '~Spare WB1[59].21'; 1910 '~Spare WB1[59].22'; 1911 '~Spare WB1[59].23'; 1912 '~Spare WB1[59].24'; 1913 '~Spare WB1[59].25'; 1914 '~Spare WB1[59].26'; 1915 '~Spare WB1[59].27'; 1916 '~Spare WB1[59].28'; 1917 '~Spare WB1[59].29'; 1918 '~Spare WB1[59].30'; 1919 '~Spare WB1[59].31'; 1920 '~S001R07 Cycle Overtime WB1[60].0'; 1921 '~S001R07 In Bypass WB1[60].1'; 1922 '~S001R07 Battery Low WB1[60].2'; 1923 '~S001R07 Servo Over Torque WB1[60].3'; 1924 '~S001R07 Process Retry In Progress WB1[60].4'; 1925 '~Spare WB1[60].5'; 1926 '~S001R07 Robot Edit Occurred Ext App WB1[60].6'; 1927 '~S001R07 Robot Input Simmed WB1[60].7'; 1928 '~S001R07 Robot Output Simmed WB1[60].8'; 1929 '~Spare WB1[60].9'; 1930 '~Spare WB1[60].10'; 1931 '~Spare WB1[60].11'; 1932 '~Spare WB1[60].12'; 1933 '~Spare WB1[60].13'; 1934 '~Spare WB1[60].14'; 1935 '~Spare WB1[60].15'; 1936 '~S001R07F1B1.M.ModuleFlt - Externa App 1 I/O Module Warning WB1[60].16'; 1937 '~S001R07F2B1.M.ModuleFlt - Externa App 2 I/O Module Warning WB1[60].17'; 1938 '~S001R07F3B1.M.ModuleFlt - Externa App 3 I/O Module Warning WB1[60].18'; 1939 '~Spare WB1[60].19'; 1940 '~Spare WB1[60].20'; 1941 '~Spare WB1[60].21'; 1942 '~Spare WB1[60].22'; 1943 '~Spare WB1[60].23'; 1944 '~S001R07ES1 - S001R07 EtherNet Switch Port At Half Duplex WB1[60].24'; 1945 '~S001R07ES1 - S001R07 EtherNet Switch Config Changes Not Saved WB1[60].25'; 1946 '~S001R07ES1 - S001R07 EtherNet Switch Configuration Changed WB1[60].26'; 1947 '~S001R07ES1 - S001R07 EtherNet Switch Port With Excessive Errors WB1[60].27'; 1948 '~S001R07ES1 - S001R07 EtherNet Switch Port With Utilization Warning WB1[60].28'; 1949 '~S001R07ES1 - S001R07 EtherNet Switch Changes Require Reboot WB1[60].29'; 1950 '~Spare WB1[60].30'; 1951 '~Spare WB1[60].31'; 1952 '~Spare WB1[61].0'; 1953 '~Spare WB1[61].1'; 1954 '~S001R07 Servo Gun Tip Calib Request 1 WB1[61].2'; 1955 '~S001R07 I-Available Warning 1 WB1[61].3'; 1956 '~S001R07 Tip Dress Motor 1 Fault Bypassed WB1[61].4'; 1957 '~S001R07 Tip Change Notice 1 WB1[61].5'; 1958 '~S001R07 Bypass Tip Dresser 1 Selected WB1[61].6'; 1959 '~S001R07 Auto Tip Changer Low 1 WB1[61].7'; 1960 '~S001R07 Auto Tip Changer Empty 1 WB1[61].8'; 1961 '~S001R07 Tip Wear Ratio Warning 1 - Touch Up Tip Dress Program WB1[61].9'; 1962 '~S001R07 Stud Weld 1 Maintenance Reqd WB1[61].10'; 1963 '~S001R07 Stud Weld 1 Low Stud Warning WB1[61].11'; 1964 '~Spare WB1[61].12'; 1965 '~S001R07 Rivet 1 Low Rivet Warning WB1[61].13'; 1966 '~S001R07 Rivet 1 - Skip Once Initiated from Robot TP WB1[61].14'; 1967 '~S001R07 Rivet 1 - Skip Remaining Initiated from Robot TP WB1[61].15'; 1968 '~S001R07 Rivet 1 Preventive Maintenace Required WB1[61].16'; 1969 '~S001R07 Rivet 1 Magazine Low WB1[61].17'; 1970 '~S001R07 Tip Change 1 Bypassed WB1[61].18'; 1971 '~S001R07 Mig Weld Fluid Level Low WB1[61].19'; 1972 '~S001R07 Weld Ctrlr 1 Adaptive Mode Is Disabled WB1[61].20'; 1973 '~S001R07 Tip Cutter 1 Warning WB1[61].21'; 1974 '~S001R07 Rivet 1 Tape-Cut Required WB1[61].22'; 1975 '~S001R07 Wire Feeder Motor Over Current WB1[61].23'; 1976 '~Spare WB1[61].24'; 1977 '~S001R07 Sealer Ctrlr 1 Minor Fault WB1[61].25'; 1978 '~S001R07 Sealer Ctrlr 1 Required Rezeroing WB1[61].26'; 1979 '~S001R07 Loaded To Average WB1[61].27'; 1980 '~S001R07 Vision Process Aborted WB1[61].28'; 1981 '~S001R07 Vision System Trending WB1[61].29'; 1982 '~S001R07 Vision Out Of Tolerance WB1[61].30'; 1983 '~Spare WB1[61].31'; 1984 '~Spare WB1[62].0'; 1985 '~Spare WB1[62].1'; 1986 '~S001R07 Servo Gun Tip Calib Request 2 WB1[62].2'; 1987 '~S001R07 I-Available Warning 2 WB1[62].3'; 1988 '~S001R07 Tip Dress Motor 2 Fault Bypassed WB1[62].4'; 1989 '~S001R07 Tip Change Notice 2 WB1[62].5'; 1990 '~S001R07 Bypass Tip Dresser 2 Selected WB1[62].6'; 1991 '~S001R07 Auto Tip Changer Low 2 WB1[62].7'; 1992 '~S001R07 Auto Tip Changer Empty 2 WB1[62].8'; 1993 '~S001R07 Tip Wear Ratio Warning 2 - Touch Up Tip Dress Program WB1[62].9'; 1994 '~S001R07 Stud Weld 2 Maintenance Reqd WB1[62].10'; 1995 '~S001R07 Stud Weld 2 Low Stud Warning WB1[62].11'; 1996 '~Spare WB1[62].12'; 1997 '~S001R07 Rivet 2 Low Rivet Warning WB1[62].13'; 1998 '~S001R07 Rivet 2 - Skip Once Initiated from Robot TP WB1[62].14'; 1999 '~S001R07 Rivet 2 - Skip Remaining Initiated from Robot TP WB1[62].15'; 2000 '~S001R07 Rivet 2 Preventive Maintenace Required WB1[62].16'; 2001 '~S001R07 Rivet 2 Magazine Low WB1[62].17'; 2002 '~S001R07 Tip Change 2 Bypassed WB1[62].18'; 2003 '~S001R07 Laser Dirty Glass Warning WB1[62].19'; 2004 '~S001R07 Weld Ctrlr 2 Adaptive Mode Is Disabled WB1[62].20'; 2005 '~S001R07 Tip Cutter 2 Warning WB1[62].21'; 2006 '~S001R07 Rivet 2 Tape-Cut Required WB1[62].22'; 2007 '~S001R07 Mig Tip Nozzel Replacement Warning WB1[62].23'; 2008 '~S001R07 Mig Tip Nozzel Replacement Required WB1[62].24'; 2009 '~S001R07 Sealer Ctrlr 2 Minor Fault WB1[62].25'; 2010 '~S001R07 Sealer Ctrlr 2 Required Rezeroing WB1[62].26'; 2011 '~S001R07 Mig Barrel Replacement Warning WB1[62].27'; 2012 '~S001R07 Mig Barrel Replacement Required WB1[62].28'; 2013 '~S001R07 In Touch Up Mode WB1[62].29'; 2014 '~S001R07 Touch Up Mode Not Enabled WB1[62].30'; 2015 '~Spare WB1[62].31'; 2016 '~S001R07 Laser Controller Fault WB1[63].0'; 2017 '~S001R07 Laser Dirty Glass Warning WB1[63].1'; 2018 '~S001R07 Laser Warning WB1[63].2'; 2019 '~Spare WB1[63].3'; 2020 '~Spare WB1[63].4'; 2021 '~Spare WB1[63].5'; 2022